(* ===== HMI "HMI_RT_1" =====
system functions are stored by id; their names below are inferred from use

ScreenModuleEditorView "Table Row" 1312x52
   TextField "tfLine" at 5,1 size 216x48; Text 'Text'
      Visibility <- "interface.tfLine.animate"
      Appearance <- "interface.tfLine.animate"
   TextField "tfTime" at 1085,1 size 222x48; Text 'Text'
      Visibility <- "interface.tfTime.animate"
      Appearance <- "interface.tfTime.animate"
   TextField "tfDropZone" at 211,1 size 236x48; Text 'Text'
      Visibility <- "interface.tfDropZone.animate"
      Appearance <- "interface.tfDropZone.animate"
   TextField "tfSLPartNumber" at 445,1 size 650x48; Text 'Text'
      Visibility <- "interface.tfPartNumber.animateSL"
      Appearance <- "interface.tfPartNumber.animateSL"
   Button "pbSelect" at 0,0 size 1312x52; TextOff 'Text'
      on Press: SetBit("interface.pbSelection.actuate")
      Appearance <- "interface.pbSelection.animate"
      ObjectEnable <- "interface.pbSelection.animate"
      Visibility <- "interface.pbSelection.animate"
      on Release: ResetBit("interface.pbSelection.actuate")
   Rectangle "rtBackground" at 0,0 size 1312x52
      Visibility <- "interface.rtBackground.animate"
      Appearance <- "interface.rtBackground.animate"
   TextField "tfDLPartNumber" at 445,1 size 650x48; Text 'Text'
      Visibility <- "interface.tfPartNumber.animateDL"
      Appearance <- "interface.tfPartNumber.animateDL"
*)

(* ===== HMI "HMI_RT_1" =====
system functions are stored by id; their names below are inferred from use

ScreenModuleEditorView "Station Sim" 102x228
   TextField "Station Label" at 0,0 size 102x20; Text 'Text'
      Appearance <- "Interface.stn.animate"
   Button "B7" at 0,22 size 50x50; TextOff 'Text'
      Appearance <- "Interface.btn.animate[7]"
      on Press: function_b14e0dd5("Interface.btn.actuate", 7)
   Button "B6" at 0,74 size 50x50; TextOff 'Text'
      Appearance <- "Interface.btn.animate[6]"
      on Press: function_b14e0dd5("Interface.btn.actuate", 6)
   Button "B5" at 0,126 size 50x50; TextOff 'Text'
      Appearance <- "Interface.btn.animate[5]"
      on Press: function_b14e0dd5("Interface.btn.actuate", 5)
   Button "B4" at 0,178 size 50x50; TextOff 'Text'
      Appearance <- "Interface.btn.animate[4]"
      on Press: function_b14e0dd5("Interface.btn.actuate", 4)
   Button "B3" at 52,22 size 50x50; TextOff 'Text'
      Appearance <- "Interface.btn.animate[3]"
      on Press: function_b14e0dd5("Interface.btn.actuate", 3)
   Button "B2" at 52,74 size 50x50; TextOff 'Text'
      Appearance <- "Interface.btn.animate[2]"
      on Press: function_b14e0dd5("Interface.btn.actuate", 2)
   Button "B1" at 52,126 size 50x50; TextOff 'Text'
      Appearance <- "Interface.btn.animate[1]"
      on Press: function_b14e0dd5("Interface.btn.actuate", 1)
   Button "B0" at 52,178 size 50x50; TextOff 'Text'
      Appearance <- "Interface.btn.animate[0]"
      on Press: function_b14e0dd5("Interface.btn.actuate", 0)
*)

(* ===== HMI "HMI_RT_1" =====
system functions are stored by id; their names below are inferred from use

ScreenModuleEditorView "Station Sim" 102x228
   TextField "Station Label" at 0,0 size 102x20; Text 'Text'
      Appearance <- "Interface.stn.animate"
   Button "B7" at 0,22 size 50x50; TextOff 'Text'
      on Press: function_b14e0dd5("Interface.btn.actuate", 7)
      Appearance <- "Interface.btn.animate[7]"
   Button "B6" at 0,74 size 50x50; TextOff 'Text'
      on Press: function_b14e0dd5("Interface.btn.actuate", 6)
      Appearance <- "Interface.btn.animate[6]"
   Button "B5" at 0,126 size 50x50; TextOff 'Text'
      on Press: function_b14e0dd5("Interface.btn.actuate", 5)
      Appearance <- "Interface.btn.animate[5]"
   Button "B4" at 0,178 size 50x50; TextOff 'Text'
      on Press: function_b14e0dd5("Interface.btn.actuate", 4)
      Appearance <- "Interface.btn.animate[4]"
   Button "B3" at 52,22 size 50x50; TextOff 'Text'
      on Press: function_b14e0dd5("Interface.btn.actuate", 3)
      Appearance <- "Interface.btn.animate[3]"
   Button "B2" at 52,74 size 50x50; TextOff 'Text'
      on Press: function_b14e0dd5("Interface.btn.actuate", 2)
      Appearance <- "Interface.btn.animate[2]"
   Button "B1" at 52,126 size 50x50; TextOff 'Text'
      on Press: function_b14e0dd5("Interface.btn.actuate", 1)
      Appearance <- "Interface.btn.animate[1]"
   Button "B0" at 52,178 size 50x50; TextOff 'Text'
      on Press: function_b14e0dd5("Interface.btn.actuate", 0)
      Appearance <- "Interface.btn.animate[0]"
*)

(* ===== HMI "HMI_RT_1" =====
system functions are stored by id; their names below are inferred from use

ScreenModuleEditorView "Station Sim" 106x232
   TextField "Station Label" at 2,2 size 102x20; Text 'Text'
      Appearance <- "Interface.stn.animate"
   Button "B7" at 2,24 size 50x50; TextOff 'Text'
      on Press: function_b14e0dd5("Interface.btn.actuate", 7)
      Appearance <- "Interface.btn.animate[7]"
   Button "B6" at 2,76 size 50x50; TextOff 'Text'
      on Press: function_b14e0dd5("Interface.btn.actuate", 6)
      Appearance <- "Interface.btn.animate[6]"
   Button "B5" at 2,128 size 50x50; TextOff 'Text'
      on Press: function_b14e0dd5("Interface.btn.actuate", 5)
      Appearance <- "Interface.btn.animate[5]"
   Button "B4" at 2,180 size 50x50; TextOff 'Text'
      on Press: function_b14e0dd5("Interface.btn.actuate", 4)
      Appearance <- "Interface.btn.animate[4]"
   Button "B3" at 54,24 size 50x50; TextOff 'Text'
      on Press: function_b14e0dd5("Interface.btn.actuate", 3)
      Appearance <- "Interface.btn.animate[3]"
   Button "B2" at 54,76 size 50x50; TextOff 'Text'
      on Press: function_b14e0dd5("Interface.btn.actuate", 2)
      Appearance <- "Interface.btn.animate[2]"
   Button "B1" at 54,128 size 50x50; TextOff 'Text'
      on Press: function_b14e0dd5("Interface.btn.actuate", 1)
      Appearance <- "Interface.btn.animate[1]"
   Button "B0" at 54,180 size 50x50; TextOff 'Text'
      on Press: function_b14e0dd5("Interface.btn.actuate", 0)
      Appearance <- "Interface.btn.animate[0]"
*)

(* ===== HMI "HMI_RT_1" =====
system functions are stored by id; their names below are inferred from use

ScreenModuleEditorView "Station Sim" 106x232
   Button "B7" at 3,26 size 48x48; TextOff 'Text'
      on Press: function_b14e0dd5("Interface.btn.actuate", 7)
      Appearance <- "Interface.btn.animate[7]"
   Button "B3" at 54,26 size 48x48; TextOff 'Text'
      on Press: function_b14e0dd5("Interface.btn.actuate", 3)
      Appearance <- "Interface.btn.animate[3]"
   Button "B6" at 3,77 size 48x48; TextOff 'Text'
      on Press: function_b14e0dd5("Interface.btn.actuate", 6)
      Appearance <- "Interface.btn.animate[6]"
   Button "B2" at 54,77 size 48x48; TextOff 'Text'
      on Press: function_b14e0dd5("Interface.btn.actuate", 2)
      Appearance <- "Interface.btn.animate[2]"
   Button "B5" at 3,128 size 48x48; TextOff 'Text'
      on Press: function_b14e0dd5("Interface.btn.actuate", 5)
      Appearance <- "Interface.btn.animate[5]"
   Button "B1" at 54,128 size 48x48; TextOff 'Text'
      on Press: function_b14e0dd5("Interface.btn.actuate", 1)
      Appearance <- "Interface.btn.animate[1]"
   Button "B4" at 3,179 size 48x48; TextOff 'Text'
      on Press: function_b14e0dd5("Interface.btn.actuate", 4)
      Appearance <- "Interface.btn.animate[4]"
   Button "B0" at 54,179 size 48x48; TextOff 'Text'
      on Press: function_b14e0dd5("Interface.btn.actuate", 0)
      Appearance <- "Interface.btn.animate[0]"
   TextField "Station Label" at 1,1 size 104x21; Text 'Text'
      Appearance <- "Interface.stn.animate"
*)

(* ===== HMI "HMI_RT_1" =====
system functions are stored by id; their names below are inferred from use

ScreenModuleEditorView "Station Sim" 106x232
   Button "B7" at 3,26 size 48x48; TextOff 'Text'
      on Press: function_b14e0dd5("Interface.btn.actuate", 7)
      Appearance <- "Interface.btn.animate[7]"
   Button "B3" at 54,26 size 48x48; TextOff 'Text'
      on Press: function_b14e0dd5("Interface.btn.actuate", 3)
      Appearance <- "Interface.btn.animate[3]"
   Button "B6" at 3,77 size 48x48; TextOff 'Text'
      on Press: function_b14e0dd5("Interface.btn.actuate", 6)
      Appearance <- "Interface.btn.animate[6]"
   Button "B2" at 54,77 size 48x48; TextOff 'Text'
      on Press: function_b14e0dd5("Interface.btn.actuate", 2)
      Appearance <- "Interface.btn.animate[2]"
   Button "B5" at 3,128 size 48x48; TextOff 'Text'
      on Press: function_b14e0dd5("Interface.btn.actuate", 5)
      Appearance <- "Interface.btn.animate[5]"
   Button "B1" at 54,128 size 48x48; TextOff 'Text'
      on Press: function_b14e0dd5("Interface.btn.actuate", 1)
      Appearance <- "Interface.btn.animate[1]"
   Button "B4" at 3,179 size 48x48; TextOff 'Text'
      on Press: function_b14e0dd5("Interface.btn.actuate", 4)
      Appearance <- "Interface.btn.animate[4]"
   Button "B0" at 54,179 size 48x48; TextOff 'Text'
      on Press: function_b14e0dd5("Interface.btn.actuate", 0)
      Appearance <- "Interface.btn.animate[0]"
   TextField "Station Label" at 1,1 size 104x21; Text 'Text'
      Appearance <- "Interface.stn.animate"
*)

(* ===== HMI "HMI_RT_1" =====
system functions are stored by id; their names below are inferred from use

ScreenModuleEditorView "Table Row" 1312x52
   TextField "tfLine" at 5,1 size 216x48; Text 'Text'
      Visibility <- "interface.tfLine.animate"
      Appearance <- "interface.tfLine.animate"
   TextField "tfTime" at 1085,1 size 222x48; Text 'Text'
      Visibility <- "interface.tfTime.animate"
      Appearance <- "interface.tfTime.animate"
   TextField "tfDropZone" at 211,1 size 236x48; Text 'Text'
      Visibility <- "interface.tfDropZone.animate"
      Appearance <- "interface.tfDropZone.animate"
   TextField "tfSLPartNumber" at 445,1 size 650x48; Text 'Text'
      Visibility <- "interface.tfPartNumber.animateSL"
      Appearance <- "interface.tfPartNumber.animateSL"
   Button "pbSelect" at 0,0 size 1312x52; TextOff 'Text'
      on Release: ResetBit("interface.pbSelection.actuate")
      on Press: SetBit("interface.pbSelection.actuate")
      Appearance <- "interface.pbSelection.animate"
      ObjectEnable <- "interface.pbSelection.animate"
      Visibility <- "interface.pbSelection.animate"
   Rectangle "rtBackground" at 0,0 size 1312x52
      Visibility <- "interface.rtBackground.animate"
      Appearance <- "interface.rtBackground.animate"
   TextField "tfDLPartNumber" at 445,1 size 650x48; Text 'Text'
      Visibility <- "interface.tfPartNumber.animateDL"
      Appearance <- "interface.tfPartNumber.animateDL"
*)

(* ===== HMI "HMI_RT_1" =====
system functions are stored by id; their names below are inferred from use

ScreenModuleEditorView "Station Assignment: Button Details" 513x74
   TextField "Button Label" at 0,0 size 75x74; Text 'Text'
      Visibility <- "Interface.label.animate"
      Appearance <- "Interface.label.animate"
   TextField "Critical Time" at 70,37 size 122x37; Text 'Text'
      Visibility <- "Interface.critical.animate"
      Appearance <- "Interface.critical.animate"
   TextField "Alloted Time" at 70,0 size 122x38; Text 'Text'
      Visibility <- "Interface.alloted.animate"
      Appearance <- "Interface.alloted.animate"
   TextField "Part Number" at 185,0 size 328x74; Text 'Text'
      Visibility <- "Interface.partNumber.animate"
      Appearance <- "Interface.partNumber.animate"
   Button "Select PB" at 0,0 size 513x74; TextOff 'Text'
      on Press: function_b14e0dd5("Interface.select.actuate", 0)
      Visibility <- "Interface.select.animate"
      ObjectEnable <- "Interface.select.animate"
*)

(* ===== HMI "HMI_RT_1" =====
system functions are stored by id; their names below are inferred from use

ScreenModuleEditorView "PB: Static Text Label" 274x45
   Button "Select All Stations" at 0,0 size 274x45; TextOff 'Text'
      on Press: function_b14e0dd5("Interface.actuate", 0)
      Appearance <- "Interface.animate"
      ObjectEnable <- "Interface.animate"
      Visibility <- "Interface.animate"
*)

(* ===== HMI "HMI_RT_1" =====
system functions are stored by id; their names below are inferred from use

ScreenModuleEditorView "PB: Station Select (Text Label)" 205x65
   Button "Station Select" at 0,0 size 205x65; TextOff 'Text'
      on Press: function_b14e0dd5("Interface.actuate", 0)
      Appearance <- "Interface.animate"
      ObjectEnable <- "Interface.animate"
      Visibility <- "Interface.animate"
*)

(* ===== HMI "HMI_RT_1" =====

ScreenModuleEditorView "PB: KP8 Stop Runtime (Text Label)" 68x66
   Button "Station Select" at 0,0 size 68x66; TextOff 'STOP RUNTIME'
      Appearance <- "Interface.animate"
      ObjectEnable <- "Interface.animate"
      Visibility <- "Interface.animate"
*)

(* ===== HMI "HMI_RT_1" =====
system functions are stored by id; their names below are inferred from use

ScreenModuleEditorView "PB: KP8 Reset Button (Text Label" 68x66
   Button "Station Select" at 0,0 size 68x66; TextOff 'RESET SELECTED'
      on Press: function_b14e0dd5("Interface.actuate", 0)
      Appearance <- "Interface.animate"
      ObjectEnable <- "Interface.animate"
      Visibility <- "Interface.animate"
*)

(* ===== HMI "HMI_RT_1" =====
system functions are stored by id; their names below are inferred from use

ScreenModuleEditorView "PB: KP8 Button Select (Text Label)" 68x66
   Button "Station Select" at 0,0 size 68x66; TextOff 'Text'
      on Press: function_b14e0dd5("Interface.actuate", 0)
      Appearance <- "Interface.animate"
      ObjectEnable <- "Interface.animate"
      Visibility <- "Interface.animate"
*)

(* ===== HMI "HMI_RT_1" =====
system functions are stored by id; their names below are inferred from use

ScreenModuleEditorView "PB: Graphic/Text List" 65x45
   Button "Previous Station Group" at 0,0 size 65x45; TextOff 'Text'
      on Press: function_b14e0dd5("Interface.actuate", 0)
      Visibility <- "Interface.animate"
      ObjectEnable <- "Interface.animate"
      Appearance <- "Interface.animate"
*)

(* ===== HMI "HMI_RT_1" =====
system functions are stored by id; their names below are inferred from use

ScreenModuleEditorView "Line Label" 267x40
   IOField "Line" at 86,0 size 181x40; FormatPattern ?????????
      on OnFinishInput: SetBit("interface.inputFinished")
      Appearance <- "interface.animate.ioField"
      Visibility <- "interface.animate.ioField"
      ObjectEnable <- "interface.animate.ioField"
      ProcessValue <- "interface.value"
   TextField "Line Label" at 0,0 size 267x40; Text 'Line:'
      Visibility <- "interface.animate.bg"
      Appearance <- "interface.animate.bg"
*)

(* ===== HMI "HMI_RT_1" =====

ScreenModuleEditorView "LED Row" 440x28
   TextField "tfLine" at 0,0 size 110x28; Text 'Text'
      Visibility <- "interface.tfLine.animate"
      Appearance <- "interface.tfLine.animate"
   TextField "tfTime" at 349,0 size 91x28; Text 'Text'
      Visibility <- "interface.tfTime.animate"
      Appearance <- "interface.tfTime.animate"
   TextField "tfDropZone" at 105,0 size 42x28; Text 'Text'
      Visibility <- "interface.tfDropZone.animate"
      Appearance <- "interface.tfDropZone.animate"
   TextField "tfSLPartNumber" at 146,0 size 209x28; Text 'Text'
      Visibility <- "interface.tfPartNumber.animateSL"
      Appearance <- "interface.tfPartNumber.animateSL"
   TextField "tfDLPartNumber" at 146,0 size 209x28; Text 'Text'
      Visibility <- "interface.tfPartNumber.animateDL"
      Appearance <- "interface.tfPartNumber.animateDL"
*)

(* ===== HMI "HMI_RT_1" =====
system functions are stored by id; their names below are inferred from use

ScreenModuleEditorView "IO Field: Timer" 137x50
   IOField "Allotted Time Entry Field" at 0,0 size 137x50; FormatPattern ???????
      on OnFinishInput: SetBit("Interface.inputFinished")
      Appearance <- "Interface.animate"
      Visibility <- "Interface.animate"
      ObjectEnable <- "Interface.animate"
      ProcessValue <- "Interface.value"
*)

(* ===== HMI "HMI_RT_1" =====
system functions are stored by id; their names below are inferred from use

ScreenModuleEditorView "IO Field: Double Width: Stacked" 414x50
   IOField "PN Entry Field" at 0,0 size 414x50; FormatPattern ????????????????????????????????????????
      on OnFinishInput: SetBit("Interface.inputFinished")
      Appearance <- "Interface.animate"
      Visibility <- "Interface.animate"
      ObjectEnable <- "Interface.animate"
      ProcessValue <- "Interface.value"
*)

(* ===== HMI "HMI_RT_1" =====
system functions are stored by id; their names below are inferred from use

ScreenModuleEditorView "Drop Zone Label" 240x40
   IOField "Drop Zone Entry" at 171,0 size 69x40; FormatPattern ??
      on OnFinishInput: SetBit("Interface.inputFinished")
      Appearance <- "Interface.animate.ioField"
      Visibility <- "Interface.animate.ioField"
      ProcessValue <- "Interface.value"
      ObjectEnable <- "Interface.animate.ioField"
   TextField "Drop Zone Label" at 0,0 size 240x40; Text 'Drop Zone:'
      Visibility <- "Interface.animate.bg"
      Appearance <- "Interface.animate.bg"
*)

(* ===== HMI "HMI_RT_1" =====
system functions are stored by id; their names below are inferred from use

ScreenModuleEditorView "PB: Station Comm Status (Text Label)" 205x65
   Button "Station Select" at 0,0 size 205x65; TextOff 'Text'
      on Press: function_b14e0dd5("Interface.actuate", 0)
      Appearance <- "Interface.animate"
      ObjectEnable <- "Interface.animate"
      Visibility <- "Interface.animate"
*)

(* ===== HMI "HMI_RT_1" =====
system functions are stored by id; their names below are inferred from use

ScreenModuleEditorView "PB: Station Comm Status (Text Label)" 180x25
   Button "Station Select" at 0,0 size 180x25; TextOff 'Text'
      on Press: function_b14e0dd5("Interface.actuate", 0)
      Appearance <- "Interface.animate"
      ObjectEnable <- "Interface.animate"
      Visibility <- "Interface.animate"
*)

(* ===== HMI "HMI_RT_1" =====
system functions are stored by id; their names below are inferred from use

ScreenModuleEditorView "PB: Station Comm Status (Text Label)" 180x25
   Button "Station Select" at 0,0 size 180x25; TextOff 'Text'
      on Press: function_b14e0dd5("Interface.actuate", 0)
      Appearance <- "Interface.animate"
      ObjectEnable <- "Interface.animate"
      Visibility <- "Interface.animate"
*)

(* ===== HMI "HMI_RT_1" =====

ScreenModuleEditorView "Station: ET200SP" 593x650
   GraphicView "ET200SP Stencil" at 0,0 size 593x649; Picture "ET 200SP Stencil"
   Rectangle "Interface Module Color" at 0,0 size 269x648
      Appearance <- "Interface.IM.bg"
   Rectangle "DQ 01 Module Color" at 268,0 size 95x342
      Appearance <- "Interface.DQ01.bg"
   Rectangle "DQ 01 Terminal Color" at 268,341 size 96x269
      Appearance <- "Interface.DQ01.bgTem"
   Rectangle "DQ 02 Module Color" at 363,1 size 96x341
      Appearance <- "Interface.DQ02.bg"
   Rectangle "DQ 02 Terminal Color" at 364,342 size 95x268
      Appearance <- "Interface.DQ02.bgTem"
   Rectangle "DQ 03 Module Color" at 458,1 size 95x342
      Appearance <- "Interface.DQ03.bg"
   Rectangle "DQ 03 Terminal Color" at 458,342 size 95x268
      Appearance <- "Interface.DQ03.bgTem"
   Rectangle "Server Module Color" at 552,1 size 40x341
      Appearance <- "Interface.serverModule.bg"
   Rectangle "IM Run LED" at 165,52 size 9x8
      Appearance <- "Interface.IM.run"
   Rectangle "IM Error LED" at 178,52 size 9x8
      Appearance <- "Interface.IM.error"
   Rectangle "IM Maintenance LED" at 193,52 size 9x8
      Appearance <- "Interface.IM.maint"
   Rectangle "IM Link 1 LED" at 146,245 size 9x8
      Appearance <- "Interface.IM.lnk01"
   Rectangle "IM Link 2 LED" at 146,263 size 9x8
      Appearance <- "Interface.IM.lnk02"
   Rectangle "IM Power LED" at 164,329 size 9x8
      Appearance <- "Interface.IM.pwr"
   Rectangle "DQ 01 Diag LED" at 274,52 size 9x8
      Appearance <- "Interface.DQ01.diag"
   Rectangle "DQ 01 Output LED x.0" at 274,245 size 9x8
      Appearance <- "Interface.DQ01.x0"
   Rectangle "DQ 01 Output LED x.1" at 305,245 size 9x8
      Appearance <- "Interface.DQ01.x1"
   Rectangle "DQ 01 Output LED x.2" at 274,256 size 9x8
      Appearance <- "Interface.DQ01.x2"
   Rectangle "DQ 01 Output LED x.3" at 305,256 size 9x8
      Appearance <- "Interface.DQ01.x3"
   Rectangle "DQ 01 Output LED x.4" at 274,267 size 9x8
      Appearance <- "Interface.DQ01.x4"
   Rectangle "DQ 01 Output LED x.5" at 305,267 size 9x8
      Appearance <- "Interface.DQ01.x5"
   Rectangle "DQ 01 Output LED x.6" at 274,278 size 9x8
      Appearance <- "Interface.DQ01.x6"
   Rectangle "DQ 01 Output LED x.7" at 305,278 size 9x8
      Appearance <- "Interface.DQ01.x7"
   Rectangle "DQ 01 Power LED" at 275,329 size 9x8
      Appearance <- "Interface.DQ01.pwr"
   Rectangle "DQ 02 Diag LED" at 369,52 size 9x8
      Appearance <- "Interface.DQ02.diag"
   Rectangle "DQ 02 Output LED x.0" at 369,245 size 9x8
      Appearance <- "Interface.DQ02.x0"
   Rectangle "DQ 02 Output LED x.1" at 400,245 size 9x8
      Appearance <- "Interface.DQ02.x1"
   Rectangle "DQ 02 Output LED x.2" at 369,256 size 9x8
      Appearance <- "Interface.DQ02.x2"
   Rectangle "DQ 02 Output LED x.3" at 400,256 size 9x8
      Appearance <- "Interface.DQ02.x3"
   Rectangle "DQ 02 Output LED x.4" at 369,267 size 9x8
      Appearance <- "Interface.DQ02.x4"
   Rectangle "DQ 02 Output LED x.5" at 400,267 size 9x8
      Appearance <- "Interface.DQ02.x5"
   Rectangle "DQ 02 Output LED x.6" at 369,278 size 9x8
      Appearance <- "Interface.DQ02.x6"
   Rectangle "DQ 02 Output LED x.7" at 400,278 size 9x8
      Appearance <- "Interface.DQ02.x7"
   Rectangle "DQ 02 Power LED" at 368,329 size 9x8
      Appearance <- "Interface.DQ02.pwr"
   Rectangle "DQ 03 Diag LED" at 464,51 size 9x8
      Appearance <- "Interface.DQ03.diag"
   Rectangle "DQ 03 Output LED x.5" at 495,267 size 9x8
      Appearance <- "Interface.DQ03.x5"
   Rectangle "DQ 03 Output LED x.6" at 464,278 size 9x8
      Appearance <- "Interface.DQ03.x6"
   Rectangle "DQ 03 Output LED x.7" at 495,278 size 9x8
      Appearance <- "Interface.DQ03.x7"
   Rectangle "DQ 03 Power LED" at 463,328 size 9x8
      Appearance <- "Interface.DQ03.pwr"
   Button "Dismiss PB" at 0,0 size 593x649; TextOff 'Text'
*)

(* ===== HMI "HMI_RT_1" =====

ScreenModuleEditorView "Station: ET200SP" 593x650
   GraphicView "ET200SP Stencil" at 0,0 size 593x649; Picture "ET 200SP Stencil"
   Rectangle "Interface Module Color" at 0,0 size 269x648
      Appearance <- "Interface.IM.bg"
   Rectangle "DQ 01 Module Color" at 268,0 size 95x342
      Appearance <- "Interface.DQ01.bg"
   Rectangle "DQ 01 Terminal Color" at 268,341 size 96x269
      Appearance <- "Interface.DQ01.bgTem"
   Rectangle "DQ 02 Module Color" at 363,1 size 96x341
      Appearance <- "Interface.DQ02.bg"
   Rectangle "DQ 02 Terminal Color" at 364,342 size 95x268
      Appearance <- "Interface.DQ02.bgTem"
   Rectangle "DQ 03 Module Color" at 458,1 size 95x342
      Appearance <- "Interface.DQ03.bg"
   Rectangle "DQ 03 Terminal Color" at 458,342 size 95x268
      Appearance <- "Interface.DQ03.bgTem"
   Rectangle "Server Module Color" at 552,1 size 40x341
      Appearance <- "Interface.serverModule.bg"
   Rectangle "IM Run LED" at 165,52 size 9x8
      Appearance <- "Interface.IM.run"
   Rectangle "IM Error LED" at 178,52 size 9x8
      Appearance <- "Interface.IM.error"
   Rectangle "IM Maintenance LED" at 193,52 size 9x8
      Appearance <- "Interface.IM.maint"
   Rectangle "IM Link 1 LED" at 146,245 size 9x8
      Appearance <- "Interface.IM.lnk01"
   Rectangle "IM Link 2 LED" at 146,263 size 9x8
      Appearance <- "Interface.IM.lnk02"
   Rectangle "IM Power LED" at 164,329 size 9x8
      Appearance <- "Interface.IM.pwr"
   Rectangle "DQ 01 Diag LED" at 274,52 size 9x8
      Appearance <- "Interface.DQ01.diag"
   Rectangle "DQ 01 Output LED x.0" at 274,245 size 9x8
      Appearance <- "Interface.DQ01.x0"
   Rectangle "DQ 01 Output LED x.1" at 305,245 size 9x8
      Appearance <- "Interface.DQ01.x1"
   Rectangle "DQ 01 Output LED x.2" at 274,256 size 9x8
      Appearance <- "Interface.DQ01.x2"
   Rectangle "DQ 01 Output LED x.3" at 305,256 size 9x8
      Appearance <- "Interface.DQ01.x3"
   Rectangle "DQ 01 Output LED x.4" at 274,267 size 9x8
      Appearance <- "Interface.DQ01.x4"
   Rectangle "DQ 01 Output LED x.5" at 305,267 size 9x8
      Appearance <- "Interface.DQ01.x5"
   Rectangle "DQ 01 Output LED x.6" at 274,278 size 9x8
      Appearance <- "Interface.DQ01.x6"
   Rectangle "DQ 01 Output LED x.7" at 305,278 size 9x8
      Appearance <- "Interface.DQ01.x7"
   Rectangle "DQ 01 Power LED" at 275,329 size 9x8
      Appearance <- "Interface.DQ01.pwr"
   Rectangle "DQ 02 Diag LED" at 369,52 size 9x8
      Appearance <- "Interface.DQ02.diag"
   Rectangle "DQ 02 Output LED x.0" at 369,245 size 9x8
      Appearance <- "Interface.DQ02.x0"
   Rectangle "DQ 02 Output LED x.1" at 400,245 size 9x8
      Appearance <- "Interface.DQ02.x1"
   Rectangle "DQ 02 Output LED x.2" at 369,256 size 9x8
      Appearance <- "Interface.DQ02.x2"
   Rectangle "DQ 02 Output LED x.3" at 400,256 size 9x8
      Appearance <- "Interface.DQ02.x3"
   Rectangle "DQ 02 Output LED x.4" at 369,267 size 9x8
      Appearance <- "Interface.DQ02.x4"
   Rectangle "DQ 02 Output LED x.5" at 400,267 size 9x8
      Appearance <- "Interface.DQ02.x5"
   Rectangle "DQ 02 Output LED x.6" at 369,278 size 9x8
      Appearance <- "Interface.DQ02.x6"
   Rectangle "DQ 02 Output LED x.7" at 400,278 size 9x8
      Appearance <- "Interface.DQ02.x7"
   Rectangle "DQ 02 Power LED" at 368,329 size 9x8
      Appearance <- "Interface.DQ02.pwr"
   Rectangle "DQ 03 Diag LED" at 464,51 size 9x8
      Appearance <- "Interface.DQ03.diag"
   Rectangle "DQ 03 Output LED x.0" at 464,245 size 9x8
      Appearance <- "Interface.DQ03.x0"
   Rectangle "DQ 03 Output LED x.1" at 495,245 size 9x8
      Appearance <- "Interface.DQ03.x1"
   Rectangle "DQ 03 Output LED x.2" at 464,256 size 9x8
      Appearance <- "Interface.DQ03.x2"
   Rectangle "DQ 03 Output LED x.3" at 495,256 size 9x8
      Appearance <- "Interface.DQ03.x3"
   Rectangle "DQ 03 Output LED x.4" at 464,267 size 9x8
      Appearance <- "Interface.DQ03.x4"
   Rectangle "DQ 03 Output LED x.5" at 495,267 size 9x8
      Appearance <- "Interface.DQ03.x5"
   Rectangle "DQ 03 Output LED x.6" at 464,278 size 9x8
      Appearance <- "Interface.DQ03.x6"
   Rectangle "DQ 03 Output LED x.7" at 495,278 size 9x8
      Appearance <- "Interface.DQ03.x7"
   Rectangle "DQ 03 Power LED" at 463,328 size 9x8
      Appearance <- "Interface.DQ03.pwr"
   Button "Dismiss PB" at 0,0 size 593x649; TextOff 'Text'
*)

(* ===== HMI "HMI_RT_1" =====

ScreenModuleEditorView "Station: ET200SP" 593x700
   GraphicView "ET200SP Stencil" at 0,50 size 593x649; Picture "ET 200SP Stencil"
   Rectangle "Interface Module Color" at 0,50 size 269x650
      Appearance <- "Interface.IM.bg"
   Rectangle "DQ 01 Module Color" at 268,50 size 95x344
      Appearance <- "Interface.DQ01.bg"
   Rectangle "DQ 01 Terminal Color" at 268,390 size 96x271
      Appearance <- "Interface.DQ01.bgTem"
   Rectangle "DQ 02 Module Color" at 363,50 size 96x344
      Appearance <- "Interface.DQ02.bg"
   Rectangle "DQ 02 Terminal Color" at 364,390 size 95x271
      Appearance <- "Interface.DQ02.bgTem"
   Rectangle "DQ 03 Module Color" at 458,50 size 95x344
      Appearance <- "Interface.DQ03.bg"
   Rectangle "DQ 03 Terminal Color" at 458,390 size 95x271
      Appearance <- "Interface.DQ03.bgTem"
   Rectangle "Server Module Color" at 552,50 size 40x343
      Appearance <- "Interface.serverModule.bg"
   Rectangle "IM Run LED" at 165,102 size 9x8
      Appearance <- "Interface.IM.run"
   Rectangle "IM Error LED" at 178,102 size 9x8
      Appearance <- "Interface.IM.error"
   Rectangle "IM Maintenance LED" at 193,102 size 9x8
      Appearance <- "Interface.IM.maint"
   Rectangle "IM Link 1 LED" at 146,295 size 9x8
      Appearance <- "Interface.IM.lnk01"
   Rectangle "IM Link 2 LED" at 146,313 size 9x8
      Appearance <- "Interface.IM.lnk02"
   Rectangle "IM Power LED" at 164,379 size 9x8
      Appearance <- "Interface.IM.pwr"
   Rectangle "DQ 01 Diag LED" at 274,102 size 9x8
      Appearance <- "Interface.DQ01.diag"
   Rectangle "DQ 01 Output LED x.0" at 274,295 size 9x8
      Appearance <- "Interface.DQ01.x0"
   Rectangle "DQ 01 Output LED x.1" at 305,295 size 9x8
      Appearance <- "Interface.DQ01.x1"
   Rectangle "DQ 01 Output LED x.2" at 274,306 size 9x8
      Appearance <- "Interface.DQ01.x2"
   Rectangle "DQ 01 Output LED x.3" at 305,306 size 9x8
      Appearance <- "Interface.DQ01.x3"
   Rectangle "DQ 01 Output LED x.4" at 274,317 size 9x8
      Appearance <- "Interface.DQ01.x4"
   Rectangle "DQ 01 Output LED x.5" at 305,317 size 9x8
      Appearance <- "Interface.DQ01.x5"
   Rectangle "DQ 01 Output LED x.6" at 274,328 size 9x8
      Appearance <- "Interface.DQ01.x6"
   Rectangle "DQ 01 Output LED x.7" at 305,328 size 9x8
      Appearance <- "Interface.DQ01.x7"
   Rectangle "DQ 01 Power LED" at 275,379 size 9x8
      Appearance <- "Interface.DQ01.pwr"
   Rectangle "DQ 02 Diag LED" at 369,102 size 9x8
      Appearance <- "Interface.DQ02.diag"
   Rectangle "DQ 02 Output LED x.0" at 369,295 size 9x8
      Appearance <- "Interface.DQ02.x0"
   Rectangle "DQ 02 Output LED x.1" at 400,295 size 9x8
      Appearance <- "Interface.DQ02.x1"
   Rectangle "DQ 02 Output LED x.2" at 369,306 size 9x8
      Appearance <- "Interface.DQ02.x2"
   Rectangle "DQ 02 Output LED x.3" at 400,306 size 9x8
      Appearance <- "Interface.DQ02.x3"
   Rectangle "DQ 02 Output LED x.4" at 369,317 size 9x8
      Appearance <- "Interface.DQ02.x4"
   Rectangle "DQ 02 Output LED x.5" at 400,317 size 9x8
      Appearance <- "Interface.DQ02.x5"
   Rectangle "DQ 02 Output LED x.6" at 369,328 size 9x8
      Appearance <- "Interface.DQ02.x6"
   Rectangle "DQ 02 Output LED x.7" at 400,328 size 9x8
      Appearance <- "Interface.DQ02.x7"
   Rectangle "DQ 02 Power LED" at 368,379 size 9x8
      Appearance <- "Interface.DQ02.pwr"
   Rectangle "DQ 03 Diag LED" at 464,102 size 9x8
      Appearance <- "Interface.DQ03.diag"
   Rectangle "DQ 03 Output LED x.0" at 464,295 size 9x8
      Appearance <- "Interface.DQ03.x0"
   Rectangle "DQ 03 Output LED x.1" at 495,295 size 9x8
      Appearance <- "Interface.DQ03.x1"
   Rectangle "DQ 03 Output LED x.2" at 464,306 size 9x8
      Appearance <- "Interface.DQ03.x2"
   Rectangle "DQ 03 Output LED x.3" at 495,306 size 9x8
      Appearance <- "Interface.DQ03.x3"
   Rectangle "DQ 03 Output LED x.4" at 464,317 size 9x8
      Appearance <- "Interface.DQ03.x4"
   Rectangle "DQ 03 Output LED x.5" at 495,317 size 9x8
      Appearance <- "Interface.DQ03.x5"
   Rectangle "DQ 03 Output LED x.6" at 464,328 size 9x8
      Appearance <- "Interface.DQ03.x6"
   Rectangle "DQ 03 Output LED x.7" at 495,328 size 9x8
      Appearance <- "Interface.DQ03.x7"
   Rectangle "DQ 03 Power LED" at 463,379 size 9x8
      Appearance <- "Interface.DQ03.pwr"
   Button "Dismiss PB" at 0,0 size 593x700; TextOff 'Text'
   TextField "PN Name" at 0,0 size 593x50; Text 'Text'
      Appearance <- "Interface.profinetName.animate"
*)

(* ===== HMI "HMI_RT_1" =====

ScreenModuleEditorView "Station: ET200SP" 603x710
   Rectangle "Interface Module Color" at 5,55 size 269x650
      Appearance <- "Interface.IM.bg"
   Rectangle "DQ 01 Module Color" at 273,55 size 95x344
      Appearance <- "Interface.DQ01.bg"
   Rectangle "DQ 01 Terminal Color" at 273,395 size 96x271
      Appearance <- "Interface.DQ01.bgTem"
   Rectangle "DQ 02 Module Color" at 368,55 size 96x344
      Appearance <- "Interface.DQ02.bg"
   Rectangle "DQ 02 Terminal Color" at 369,395 size 95x271
      Appearance <- "Interface.DQ02.bgTem"
   Rectangle "DQ 03 Module Color" at 463,55 size 95x344
      Appearance <- "Interface.DQ03.bg"
   Rectangle "DQ 03 Terminal Color" at 463,395 size 95x271
      Appearance <- "Interface.DQ03.bgTem"
   Rectangle "Server Module Color" at 557,55 size 40x343
      Appearance <- "Interface.serverModule.bg"
   Rectangle "IM Run LED" at 170,107 size 9x8
      Appearance <- "Interface.IM.run"
   Rectangle "IM Error LED" at 183,107 size 9x8
      Appearance <- "Interface.IM.error"
   Rectangle "IM Maintenance LED" at 198,107 size 9x8
      Appearance <- "Interface.IM.maint"
   Rectangle "IM Link 1 LED" at 151,300 size 9x8
      Appearance <- "Interface.IM.lnk01"
   Rectangle "IM Link 2 LED" at 151,318 size 9x8
      Appearance <- "Interface.IM.lnk02"
   Rectangle "IM Power LED" at 169,384 size 9x8
      Appearance <- "Interface.IM.pwr"
   Rectangle "DQ 01 Diag LED" at 279,107 size 9x8
      Appearance <- "Interface.DQ01.diag"
   Rectangle "DQ 01 Output LED x.0" at 279,300 size 9x8
      Appearance <- "Interface.DQ01.x0"
   Rectangle "DQ 01 Output LED x.1" at 310,300 size 9x8
      Appearance <- "Interface.DQ01.x1"
   Rectangle "DQ 01 Output LED x.2" at 279,311 size 9x8
      Appearance <- "Interface.DQ01.x2"
   Rectangle "DQ 01 Output LED x.3" at 310,311 size 9x8
      Appearance <- "Interface.DQ01.x3"
   Rectangle "DQ 01 Output LED x.4" at 279,322 size 9x8
      Appearance <- "Interface.DQ01.x4"
   Rectangle "DQ 01 Output LED x.5" at 310,322 size 9x8
      Appearance <- "Interface.DQ01.x5"
   Rectangle "DQ 01 Output LED x.6" at 279,333 size 9x8
      Appearance <- "Interface.DQ01.x6"
   Rectangle "DQ 01 Output LED x.7" at 310,333 size 9x8
      Appearance <- "Interface.DQ01.x7"
   Rectangle "DQ 01 Power LED" at 280,384 size 9x8
      Appearance <- "Interface.DQ01.pwr"
   Rectangle "DQ 02 Diag LED" at 374,107 size 9x8
      Appearance <- "Interface.DQ02.diag"
   Rectangle "DQ 02 Output LED x.0" at 374,300 size 9x8
      Appearance <- "Interface.DQ02.x0"
   Rectangle "DQ 02 Output LED x.1" at 405,300 size 9x8
      Appearance <- "Interface.DQ02.x1"
   Rectangle "DQ 02 Output LED x.2" at 374,311 size 9x8
      Appearance <- "Interface.DQ02.x2"
   Rectangle "DQ 02 Output LED x.3" at 405,311 size 9x8
      Appearance <- "Interface.DQ02.x3"
   Rectangle "DQ 02 Output LED x.4" at 374,322 size 9x8
      Appearance <- "Interface.DQ02.x4"
   Rectangle "DQ 02 Output LED x.5" at 405,322 size 9x8
      Appearance <- "Interface.DQ02.x5"
   Rectangle "DQ 02 Output LED x.6" at 374,333 size 9x8
      Appearance <- "Interface.DQ02.x6"
   Rectangle "DQ 02 Output LED x.7" at 405,333 size 9x8
      Appearance <- "Interface.DQ02.x7"
   Rectangle "DQ 02 Power LED" at 373,384 size 9x8
      Appearance <- "Interface.DQ02.pwr"
   Rectangle "DQ 03 Diag LED" at 469,107 size 9x8
      Appearance <- "Interface.DQ03.diag"
   Rectangle "DQ 03 Output LED x.0" at 469,300 size 9x8
      Appearance <- "Interface.DQ03.x0"
   Rectangle "DQ 03 Output LED x.1" at 500,300 size 9x8
      Appearance <- "Interface.DQ03.x1"
   Rectangle "DQ 03 Output LED x.2" at 469,311 size 9x8
      Appearance <- "Interface.DQ03.x2"
   Rectangle "DQ 03 Output LED x.3" at 500,311 size 9x8
      Appearance <- "Interface.DQ03.x3"
   Rectangle "DQ 03 Output LED x.4" at 469,322 size 9x8
      Appearance <- "Interface.DQ03.x4"
   Rectangle "DQ 03 Output LED x.5" at 500,322 size 9x8
      Appearance <- "Interface.DQ03.x5"
   Rectangle "DQ 03 Output LED x.6" at 469,333 size 9x8
      Appearance <- "Interface.DQ03.x6"
   Rectangle "DQ 03 Output LED x.7" at 500,333 size 9x8
      Appearance <- "Interface.DQ03.x7"
   Rectangle "DQ 03 Power LED" at 468,384 size 9x8
      Appearance <- "Interface.DQ03.pwr"
   GraphicView "ET200SP Stencil" at 5,55 size 593x649; Picture "ET 200SP Stencil"
   Button "Dismiss PB" at 5,5 size 593x700; TextOff 'Text'
   TextField "PN Name" at 5,5 size 593x50; Text 'Text'
      Appearance <- "Interface.profinetName.animate"
*)

(* ===== HMI "HMI_RT_1" =====

ScreenModuleEditorView "Station: KP8" 428x710
   GraphicView "KP8 Stencil" at 5,55 size 418x650; Picture "KP8 Rear View Stencil"
      Appearance <- "Interface.stencilBackground"
   TextField "PN Name Label" at 5,5 size 418x50; Text 'Text'
      Appearance <- "Interface.profinetName.animate"
   Rectangle "X1P1 Transmit" at 195,536 size 12x16
      Appearance <- "Interface.X1P1.transmit"
   Rectangle "X1P1 Receive" at 195,576 size 12x16
      Appearance <- "Interface.X1P1.receive"
   Rectangle "X1P2 Transmit" at 286,535 size 12x16
      Appearance <- "Interface.X1P2.transmit"
   Rectangle "X1P2 Receive" at 286,575 size 12x16
      Appearance <- "Interface.X1P2.receive"
   Rectangle "KP8 Background" at 5,55 size 418x650
      Appearance <- "Interface.profinetName.animate"
   Button "Dissmiss PB" at 5,5 size 418x700; TextOff 'Text'
*)

(* ===== HMI "HMI_RT_1" =====

ScreenModuleEditorView "Station: ET200SP" 603x710
   TextField "PN Name" at 5,5 size 593x50; Text 'Text'
      Appearance <- "Interface.profinetName.animate"
   Rectangle "Interface Module Color" at 5,55 size 269x650
      Appearance <- "Interface.IM.bg"
   Rectangle "DQ 01 Module Color" at 273,55 size 95x344
      Appearance <- "Interface.DQ01.bg"
   Rectangle "DQ 01 Terminal Color" at 273,395 size 96x271
      Appearance <- "Interface.DQ01.bgTem"
   Rectangle "DQ 02 Module Color" at 368,55 size 96x344
      Appearance <- "Interface.DQ02.bg"
   Rectangle "DQ 02 Terminal Color" at 369,395 size 95x271
      Appearance <- "Interface.DQ02.bgTem"
   Rectangle "DQ 03 Module Color" at 463,55 size 95x344
      Appearance <- "Interface.DQ03.bg"
   Rectangle "DQ 03 Terminal Color" at 463,395 size 95x271
      Appearance <- "Interface.DQ03.bgTem"
   Rectangle "Server Module Color" at 557,55 size 40x343
      Appearance <- "Interface.serverModule.bg"
   Rectangle "IM Run LED" at 170,107 size 9x8
      Appearance <- "Interface.IM.run"
   Rectangle "IM Error LED" at 183,107 size 9x8
      Appearance <- "Interface.IM.error"
   Rectangle "IM Maintenance LED" at 198,107 size 9x8
      Appearance <- "Interface.IM.maint"
   Rectangle "IM Link 1 LED" at 151,300 size 9x8
      Appearance <- "Interface.IM.lnk01"
   Rectangle "IM Link 2 LED" at 151,318 size 9x8
      Appearance <- "Interface.IM.lnk02"
   Rectangle "IM Power LED" at 169,384 size 9x8
      Appearance <- "Interface.IM.pwr"
   Rectangle "DQ 01 Diag LED" at 279,107 size 9x8
      Appearance <- "Interface.DQ01.diag"
   Rectangle "DQ 01 Output LED x.0" at 279,300 size 9x8
      Appearance <- "Interface.DQ01.x0"
   Rectangle "DQ 01 Output LED x.1" at 310,300 size 9x8
      Appearance <- "Interface.DQ01.x1"
   Rectangle "DQ 01 Output LED x.2" at 279,311 size 9x8
      Appearance <- "Interface.DQ01.x2"
   Rectangle "DQ 01 Output LED x.3" at 310,311 size 9x8
      Appearance <- "Interface.DQ01.x3"
   Rectangle "DQ 01 Output LED x.4" at 279,322 size 9x8
      Appearance <- "Interface.DQ01.x4"
   Rectangle "DQ 01 Output LED x.5" at 310,322 size 9x8
      Appearance <- "Interface.DQ01.x5"
   Rectangle "DQ 01 Output LED x.6" at 279,333 size 9x8
      Appearance <- "Interface.DQ01.x6"
   Rectangle "DQ 01 Output LED x.7" at 310,333 size 9x8
      Appearance <- "Interface.DQ01.x7"
   Rectangle "DQ 01 Power LED" at 280,384 size 9x8
      Appearance <- "Interface.DQ01.pwr"
   Rectangle "DQ 02 Diag LED" at 374,107 size 9x8
      Appearance <- "Interface.DQ02.diag"
   Rectangle "DQ 02 Output LED x.0" at 374,300 size 9x8
      Appearance <- "Interface.DQ02.x0"
   Rectangle "DQ 02 Output LED x.1" at 405,300 size 9x8
      Appearance <- "Interface.DQ02.x1"
   Rectangle "DQ 02 Output LED x.2" at 374,311 size 9x8
      Appearance <- "Interface.DQ02.x2"
   Rectangle "DQ 02 Output LED x.3" at 405,311 size 9x8
      Appearance <- "Interface.DQ02.x3"
   Rectangle "DQ 02 Output LED x.4" at 374,322 size 9x8
      Appearance <- "Interface.DQ02.x4"
   Rectangle "DQ 02 Output LED x.5" at 405,322 size 9x8
      Appearance <- "Interface.DQ02.x5"
   Rectangle "DQ 02 Output LED x.6" at 374,333 size 9x8
      Appearance <- "Interface.DQ02.x6"
   Rectangle "DQ 02 Output LED x.7" at 405,333 size 9x8
      Appearance <- "Interface.DQ02.x7"
   Rectangle "DQ 02 Power LED" at 373,384 size 9x8
      Appearance <- "Interface.DQ02.pwr"
   Rectangle "DQ 03 Diag LED" at 469,107 size 9x8
      Appearance <- "Interface.DQ03.diag"
   Rectangle "DQ 03 Output LED x.0" at 469,300 size 9x8
      Appearance <- "Interface.DQ03.x0"
   Rectangle "DQ 03 Output LED x.1" at 500,300 size 9x8
      Appearance <- "Interface.DQ03.x1"
   Rectangle "DQ 03 Output LED x.2" at 469,311 size 9x8
      Appearance <- "Interface.DQ03.x2"
   Rectangle "DQ 03 Output LED x.3" at 500,311 size 9x8
      Appearance <- "Interface.DQ03.x3"
   Rectangle "DQ 03 Output LED x.4" at 469,322 size 9x8
      Appearance <- "Interface.DQ03.x4"
   Rectangle "DQ 03 Output LED x.5" at 500,322 size 9x8
      Appearance <- "Interface.DQ03.x5"
   Rectangle "DQ 03 Output LED x.6" at 469,333 size 9x8
      Appearance <- "Interface.DQ03.x6"
   Rectangle "DQ 03 Output LED x.7" at 500,333 size 9x8
      Appearance <- "Interface.DQ03.x7"
   Rectangle "DQ 03 Power LED" at 468,384 size 9x8
      Appearance <- "Interface.DQ03.pwr"
   GraphicView "ET200SP Stencil" at 5,55 size 593x649; Picture "ET 200SP Stencil"
   Button "Dismiss PB" at 5,5 size 593x700; TextOff 'Text'
*)

(* ===== HMI "HMI_RT_6" =====
system functions are stored by id; their names below are inferred from use
connection "cv01": ETHERNET, SMART_S7_1500_OMS

HMI tags "Default tag table"
   "station" : HMI Station: Compressed = PLC "HMI Data: TP700 Stations".stns[0] AT %DB1.DBW0, 100 ms

screen "01 Part Select" 480x800, template "Current Menu Selection"
   Button "B7" at 6,164 size 233x154; TextOff 'Text'
      on Press: function_b14e0dd5("pbs", 7)
      Visibility <- "[7]"
   Button "B6" at 6,323 size 233x154; TextOff 'Text'
      on Press: function_b14e0dd5("pbs", 6)
      Visibility <- "[6]"
   Button "B5" at 6,482 size 233x154; TextOff 'Text'
      on Press: function_b14e0dd5("pbs", 5)
      Visibility <- "[5]"
   Button "B4" at 6,641 size 233x154; TextOff 'Text'
      on Press: function_b14e0dd5("pbs", 4)
      Visibility <- "[4]"
   Button "B3" at 244,164 size 232x154; TextOff 'Text'
      on Press: function_b14e0dd5("pbs", 3)
      Visibility <- "[3]"
   Button "B2" at 244,323 size 232x154; TextOff 'Text'
      on Press: function_b14e0dd5("pbs", 2)
      Visibility <- "[2]"
   Button "B1" at 244,482 size 232x154; TextOff 'Text'
      on Press: function_b14e0dd5("pbs", 1)
      Visibility <- "[1]"
   Button "B0" at 244,641 size 232x154; TextOff 'Text'
      on Press: function_b14e0dd5("pbs", 0)
   IOField "B7 Label" at 6,164 size 233x154; FormatPattern ????????????????????????????????????????
      Appearance <- "[7]"
      ProcessValue <- "[7]"
      Visibility <- "[7]"
   IOField "B6 Label" at 6,323 size 233x154; FormatPattern ????????????????????????????????????????
      Appearance <- "[6]"
      ProcessValue <- "[6]"
      Visibility <- "[6]"
   IOField "B5 Label" at 6,482 size 233x154; FormatPattern ????????????????????????????????????????
      Appearance <- "[5]"
      ProcessValue <- "[5]"
      Visibility <- "[5]"
   IOField "B4 Label" at 6,641 size 233x154; FormatPattern ????????????????????????????????????????
      Appearance <- "[4]"
      ProcessValue <- "[4]"
      Visibility <- "[4]"
   IOField "B3 Label" at 244,164 size 232x154; FormatPattern ????????????????????????????????????????
      Appearance <- "[3]"
      ProcessValue <- "[3]"
      Visibility <- "[3]"
   IOField "B2 Label" at 244,323 size 232x154; FormatPattern ????????????????????????????????????????
      Appearance <- "[2]"
      ProcessValue <- "[2]"
      Visibility <- "[2]"
   IOField "B1 Label" at 244,482 size 232x154; FormatPattern ????????????????????????????????????????
      Appearance <- "[1]"
      ProcessValue <- "[1]"
      Visibility <- "[1]"
   IOField "B0 Label" at 244,641 size 232x154; FormatPattern ????????????????????????????????????????
      Appearance <- "[0]"
      ProcessValue <- "[0]"
      Visibility <- "[0]"
   TextField "B7 BG" at 6,164 size 233x154; Text '1'
      Appearance <- "[7]"
      Visibility <- "[7]"
   TextField "B6 BG" at 6,323 size 233x154; Text '3'
      Appearance <- "[6]"
      Visibility <- "[6]"
   TextField "B5 BG" at 6,482 size 233x154; Text '5'
      Appearance <- "[5]"
      Visibility <- "[5]"
   TextField "B4 BG" at 6,641 size 233x154; Text '7'
      Appearance <- "[4]"
      Visibility <- "[4]"
   TextField "B3 BG" at 244,164 size 233x154; Text '2'
      Appearance <- "[3]"
      Visibility <- "[3]"
   TextField "B2 BG" at 244,323 size 233x154; Text '4'
      Appearance <- "[2]"
      Visibility <- "[2]"
   TextField "B1 BG" at 244,482 size 233x154; Text '6'
      Appearance <- "[1]"
      Visibility <- "[1]"
   TextField "B0 BG" at 244,641 size 233x154; Text '8'
      Appearance <- "[0]"
      Visibility <- "[0]"